DATA_BLOCK "DB1901_Config_Robots"   // DB1901
{ S7_Optimized_Access := 'FALSE' }
VERSION : 0.1
   VAR
      ReadWriteDeviceNo : Int := 1;
      CopyDeviceNO : Int := 0;
      Read : Bool := FALSE;
      Write : Bool := FALSE;
      Copy : Bool := FALSE;
      Config_Robots : Array[0..4] of Struct
         Type_Kuka : Bool;   // Kuka Robot
         Type_ABB : Bool;   // ABB Robot
         Type_Fanuc : Bool;   // Fanuc Robot
         Type_Motoman : Bool;   // Motoman (Yaskawa) Robot
         Type_5 : Bool;
         Type_6 : Bool;
         Type_7 : Bool;
         Type_8 : Bool;
         With_Shotware : Bool;   // Only ABB
         With_Tracking : Bool;
         With_Safetysoftware : Bool;   // EPS/Safemove or simmilar
         With_Synchronisation : Bool;   // EPS Sync switch, Breaktest, ...
         With_Testshot : Bool;   // With Test shot station
         With_Cleaning : Bool;   // With Cleaning (automaitc)
         With_Wet_Cleaning : Bool;   // With wet cleaning
         With_Wet_Cleaning_LFI : Bool;   // Water cleaning LFI
         With_Wet_Cleaning_Spray : Bool;   // Wet cleaning Spray
         With_IR_Station : Bool;   // With Infra red station
         With_Brush_Station : Bool;   // With Brush station (motor)
         With_Belt_Filter : Bool;   // With belt filter for LFI wet cleaning
         With_Air_Cleaner : Bool;   // With Air cleaning system for the mixinghead
         Spare_2_5 : Bool;
         Spare_2_6 : Bool;
         Spare_2_7 : Bool;
         MHNumber : Byte;
         InterfaceForTestShot : Byte;
         ForInterface : Array[1..16] of Bool;
      END_STRUCT;
   END_VAR
BEGIN
   Config_Robots[0].Type_Kuka := FALSE;
   Config_Robots[0].Type_ABB := FALSE;
   Config_Robots[0].Type_Fanuc := FALSE;
   Config_Robots[0].Type_Motoman := FALSE;
   Config_Robots[0].Type_5 := FALSE;
   Config_Robots[0].Type_6 := FALSE;
   Config_Robots[0].Type_7 := FALSE;
   Config_Robots[0].Type_8 := FALSE;
   Config_Robots[0].With_Shotware := FALSE;
   Config_Robots[0].With_Tracking := FALSE;
   Config_Robots[0].With_Safetysoftware := FALSE;
   Config_Robots[0].With_Synchronisation := TRUE;
   Config_Robots[0].With_Testshot := TRUE;
   Config_Robots[0].With_Cleaning := TRUE;
   Config_Robots[0].With_Wet_Cleaning := FALSE;
   Config_Robots[0].With_Wet_Cleaning_LFI := FALSE;
   Config_Robots[0].With_Wet_Cleaning_Spray := FALSE;
   Config_Robots[0].With_IR_Station := FALSE;
   Config_Robots[0].With_Brush_Station := FALSE;
   Config_Robots[0].With_Belt_Filter := FALSE;
   Config_Robots[0].With_Air_Cleaner := FALSE;
   Config_Robots[0].Spare_2_5 := FALSE;
   Config_Robots[0].Spare_2_6 := FALSE;
   Config_Robots[0].Spare_2_7 := FALSE;
   Config_Robots[1].Type_Kuka := FALSE;
   Config_Robots[1].Type_ABB := FALSE;
   Config_Robots[1].Type_Fanuc := FALSE;
   Config_Robots[1].Type_Motoman := FALSE;
   Config_Robots[1].Type_5 := FALSE;
   Config_Robots[1].Type_6 := FALSE;
   Config_Robots[1].Type_7 := FALSE;
   Config_Robots[1].Type_8 := FALSE;
   Config_Robots[1].With_Shotware := FALSE;
   Config_Robots[1].With_Tracking := FALSE;
   Config_Robots[1].With_Safetysoftware := FALSE;
   Config_Robots[1].With_Synchronisation := TRUE;
   Config_Robots[1].With_Testshot := TRUE;
   Config_Robots[1].With_Cleaning := TRUE;
   Config_Robots[1].With_Wet_Cleaning := FALSE;
   Config_Robots[1].With_Wet_Cleaning_LFI := FALSE;
   Config_Robots[1].With_Wet_Cleaning_Spray := FALSE;
   Config_Robots[1].With_IR_Station := FALSE;
   Config_Robots[1].With_Brush_Station := FALSE;
   Config_Robots[1].With_Belt_Filter := FALSE;
   Config_Robots[1].With_Air_Cleaner := FALSE;
   Config_Robots[1].Spare_2_5 := FALSE;
   Config_Robots[1].Spare_2_6 := FALSE;
   Config_Robots[1].Spare_2_7 := FALSE;
   Config_Robots[2].Type_Kuka := FALSE;
   Config_Robots[2].Type_ABB := FALSE;
   Config_Robots[2].Type_Fanuc := FALSE;
   Config_Robots[2].Type_Motoman := FALSE;
   Config_Robots[2].Type_5 := FALSE;
   Config_Robots[2].Type_6 := FALSE;
   Config_Robots[2].Type_7 := FALSE;
   Config_Robots[2].Type_8 := FALSE;
   Config_Robots[2].With_Shotware := FALSE;
   Config_Robots[2].With_Tracking := FALSE;
   Config_Robots[2].With_Safetysoftware := FALSE;
   Config_Robots[2].With_Synchronisation := FALSE;
   Config_Robots[2].With_Testshot := FALSE;
   Config_Robots[2].With_Cleaning := FALSE;
   Config_Robots[2].With_Wet_Cleaning := FALSE;
   Config_Robots[2].With_Wet_Cleaning_LFI := FALSE;
   Config_Robots[2].With_Wet_Cleaning_Spray := FALSE;
   Config_Robots[2].With_IR_Station := FALSE;
   Config_Robots[2].With_Brush_Station := FALSE;
   Config_Robots[2].With_Belt_Filter := FALSE;
   Config_Robots[2].With_Air_Cleaner := FALSE;
   Config_Robots[2].Spare_2_5 := FALSE;
   Config_Robots[2].Spare_2_6 := FALSE;
   Config_Robots[2].Spare_2_7 := FALSE;
   Config_Robots[3].Type_Kuka := FALSE;
   Config_Robots[3].Type_ABB := FALSE;
   Config_Robots[3].Type_Fanuc := FALSE;
   Config_Robots[3].Type_Motoman := FALSE;
   Config_Robots[3].Type_5 := FALSE;
   Config_Robots[3].Type_6 := FALSE;
   Config_Robots[3].Type_7 := FALSE;
   Config_Robots[3].Type_8 := FALSE;
   Config_Robots[3].With_Shotware := FALSE;
   Config_Robots[3].With_Tracking := FALSE;
   Config_Robots[3].With_Safetysoftware := FALSE;
   Config_Robots[3].With_Synchronisation := FALSE;
   Config_Robots[3].With_Testshot := FALSE;
   Config_Robots[3].With_Cleaning := FALSE;
   Config_Robots[3].With_Wet_Cleaning := FALSE;
   Config_Robots[3].With_Wet_Cleaning_LFI := FALSE;
   Config_Robots[3].With_Wet_Cleaning_Spray := FALSE;
   Config_Robots[3].With_IR_Station := FALSE;
   Config_Robots[3].With_Brush_Station := FALSE;
   Config_Robots[3].With_Belt_Filter := FALSE;
   Config_Robots[3].With_Air_Cleaner := FALSE;
   Config_Robots[3].Spare_2_5 := FALSE;
   Config_Robots[3].Spare_2_6 := FALSE;
   Config_Robots[3].Spare_2_7 := FALSE;
   Config_Robots[4].Type_Kuka := FALSE;
   Config_Robots[4].Type_ABB := FALSE;
   Config_Robots[4].Type_Fanuc := FALSE;
   Config_Robots[4].Type_Motoman := FALSE;
   Config_Robots[4].Type_5 := FALSE;
   Config_Robots[4].Type_6 := FALSE;
   Config_Robots[4].Type_7 := FALSE;
   Config_Robots[4].Type_8 := FALSE;
   Config_Robots[4].With_Shotware := FALSE;
   Config_Robots[4].With_Tracking := FALSE;
   Config_Robots[4].With_Safetysoftware := FALSE;
   Config_Robots[4].With_Synchronisation := FALSE;
   Config_Robots[4].With_Testshot := FALSE;
   Config_Robots[4].With_Cleaning := FALSE;
   Config_Robots[4].With_Wet_Cleaning := FALSE;
   Config_Robots[4].With_Wet_Cleaning_LFI := FALSE;
   Config_Robots[4].With_Wet_Cleaning_Spray := FALSE;
   Config_Robots[4].With_IR_Station := FALSE;
   Config_Robots[4].With_Brush_Station := FALSE;
   Config_Robots[4].With_Belt_Filter := FALSE;
   Config_Robots[4].With_Air_Cleaner := FALSE;
   Config_Robots[4].Spare_2_5 := FALSE;
   Config_Robots[4].Spare_2_6 := FALSE;
   Config_Robots[4].Spare_2_7 := FALSE;
   Config_Robots[1].ForInterface[1] := TRUE;
   Config_Robots[1].ForInterface[2] := TRUE;
   Config_Robots[1].ForInterface[3] := TRUE;
   Config_Robots[1].ForInterface[4] := TRUE;
   Config_Robots[1].ForInterface[5] := TRUE;
   Config_Robots[1].InterfaceForTestShot := 16#05;
   Config_Robots[0].MHNumber := 16#01;
   Config_Robots[0].InterfaceForTestShot := 16#05;
   Config_Robots[0].ForInterface[1] := TRUE;
   Config_Robots[0].ForInterface[2] := TRUE;
   Config_Robots[0].ForInterface[3] := TRUE;
   Config_Robots[0].ForInterface[4] := TRUE;
   Config_Robots[0].ForInterface[5] := TRUE;
   Config_Robots[0].ForInterface[6] := FALSE;
   Config_Robots[0].ForInterface[7] := FALSE;
   Config_Robots[0].ForInterface[8] := FALSE;
   Config_Robots[0].ForInterface[9] := FALSE;
   Config_Robots[0].ForInterface[10] := FALSE;
   Config_Robots[0].ForInterface[11] := FALSE;
   Config_Robots[0].ForInterface[12] := FALSE;
   Config_Robots[0].ForInterface[13] := FALSE;
   Config_Robots[0].ForInterface[14] := FALSE;
   Config_Robots[0].ForInterface[15] := FALSE;
   Config_Robots[0].ForInterface[16] := FALSE;
   Config_Robots[1].MHNumber := 16#01;
   Config_Robots[1].ForInterface[6] := FALSE;
   Config_Robots[1].ForInterface[7] := FALSE;
   Config_Robots[1].ForInterface[8] := FALSE;
   Config_Robots[1].ForInterface[9] := FALSE;
   Config_Robots[1].ForInterface[10] := FALSE;
   Config_Robots[1].ForInterface[11] := FALSE;
   Config_Robots[1].ForInterface[12] := FALSE;
   Config_Robots[1].ForInterface[13] := FALSE;
   Config_Robots[1].ForInterface[14] := FALSE;
   Config_Robots[1].ForInterface[15] := FALSE;
   Config_Robots[1].ForInterface[16] := FALSE;
   Config_Robots[2].MHNumber := 16#00;
   Config_Robots[2].InterfaceForTestShot := 16#00;
   Config_Robots[2].ForInterface[1] := FALSE;
   Config_Robots[2].ForInterface[2] := FALSE;
   Config_Robots[2].ForInterface[3] := FALSE;
   Config_Robots[2].ForInterface[4] := FALSE;
   Config_Robots[2].ForInterface[5] := FALSE;
   Config_Robots[2].ForInterface[6] := FALSE;
   Config_Robots[2].ForInterface[7] := FALSE;
   Config_Robots[2].ForInterface[8] := FALSE;
   Config_Robots[2].ForInterface[9] := FALSE;
   Config_Robots[2].ForInterface[10] := FALSE;
   Config_Robots[2].ForInterface[11] := FALSE;
   Config_Robots[2].ForInterface[12] := FALSE;
   Config_Robots[2].ForInterface[13] := FALSE;
   Config_Robots[2].ForInterface[14] := FALSE;
   Config_Robots[2].ForInterface[15] := FALSE;
   Config_Robots[2].ForInterface[16] := FALSE;
   Config_Robots[3].MHNumber := 16#00;
   Config_Robots[3].InterfaceForTestShot := 16#00;
   Config_Robots[3].ForInterface[1] := FALSE;
   Config_Robots[3].ForInterface[2] := FALSE;
   Config_Robots[3].ForInterface[3] := FALSE;
   Config_Robots[3].ForInterface[4] := FALSE;
   Config_Robots[3].ForInterface[5] := FALSE;
   Config_Robots[3].ForInterface[6] := FALSE;
   Config_Robots[3].ForInterface[7] := FALSE;
   Config_Robots[3].ForInterface[8] := FALSE;
   Config_Robots[3].ForInterface[9] := FALSE;
   Config_Robots[3].ForInterface[10] := FALSE;
   Config_Robots[3].ForInterface[11] := FALSE;
   Config_Robots[3].ForInterface[12] := FALSE;
   Config_Robots[3].ForInterface[13] := FALSE;
   Config_Robots[3].ForInterface[14] := FALSE;
   Config_Robots[3].ForInterface[15] := FALSE;
   Config_Robots[3].ForInterface[16] := FALSE;
   Config_Robots[4].MHNumber := 16#00;
   Config_Robots[4].InterfaceForTestShot := 16#00;
   Config_Robots[4].ForInterface[1] := FALSE;
   Config_Robots[4].ForInterface[2] := FALSE;
   Config_Robots[4].ForInterface[3] := FALSE;
   Config_Robots[4].ForInterface[4] := FALSE;
   Config_Robots[4].ForInterface[5] := FALSE;
   Config_Robots[4].ForInterface[6] := FALSE;
   // 10 more start values not shown
END_DATA_BLOCK

DATA_BLOCK "GetToolShotValues_DB"   // DB1930
{ S7_Optimized_Access := 'FALSE' }
VERSION : 0.1
"GetToolShotValues"
BEGIN
   IN_MachineNo := 1;
   IN_EnableTool := TRUE;
END_DATA_BLOCK

DATA_BLOCK "FB1931_ToolAllocationList_DB"   // DB1931
{ S7_Optimized_Access := 'TRUE' }
VERSION : 0.1
"FB1931_ToolAllocationList"
BEGIN
END_DATA_BLOCK

DATA_BLOCK "DB2000_FRA<->KM"   // DB2000
{ S7_Optimized_Access := 'FALSE' }
VERSION : 0.1
   VAR
      AP_Shottime : Int := 0;   // Schusszeit in ms
      AP_MVH : Int := 0;   // Mischungsverhältnis in 0,1%
      AP_Weight : Int := 0;   // Gesamtgewicht pro Sekunde in 0,1 Gramm
      FRA1_Stat : "UDT2000_KM_FRA";
      FRA1_PrgNr : Byte := B#16#0;
      Bit_FT1_sel : Bool := FALSE;
      Bit_FRA1_Sel : Bool := FALSE;
      TS1_Offset : Byte := B#16#0;
      Input : "UDT2001_Input_Faurecia";
      Output : "UDT2002_Output_Faurecia";
   END_VAR
BEGIN
END_DATA_BLOCK

DATA_BLOCK "PN_Devices"   // DB2023
{ S7_Optimized_Access := 'TRUE' }
VERSION : 0.1
   VAR
      LADDR : Hw_IoSystem := 257;
      MODE : UInt := 4;
      RETVAL : Int;
      Device_available : Array[0..1023] of Bool;
   END_VAR
BEGIN
   // Device_available[2] : pn-mixhead
   // Device_available[1] : pn-flow1
   // Device_available[0] : Bei mindestens einem der IO-Devices liegt eine Störung vor.
END_DATA_BLOCK

DATA_BLOCK "PB_Devices"   // DB2024
{ S7_Optimized_Access := 'TRUE' }
VERSION : 0.1
   VAR
      LADDR : Hw_IoSystem := 296;
      MODE : UInt := 4;
      RETVAL : Int;
      Device_available : Array[0..127] of Bool;
   END_VAR
BEGIN
END_DATA_BLOCK

// folder: System blocks/Program resources

DATA_BLOCK "DB55_Temp_HD_WT_MK1_K1"   // DB55
{ S7_Optimized_Access := 'TRUE' }
AUTHOR : Simatic
FAMILY : IEC
NAME : IEC_TMR
VERSION : 1.0
"IEC_TIMER"
BEGIN
END_DATA_BLOCK

DATA_BLOCK "DB56_Temp_HD_WT_MK1_K2"   // DB56
{ S7_Optimized_Access := 'TRUE' }
AUTHOR : Simatic
FAMILY : IEC
NAME : IEC_TMR
VERSION : 1.0
"IEC_TIMER"
BEGIN
END_DATA_BLOCK

DATA_BLOCK "DB60_Temp_ND_WT_MK1_K1"   // DB60
{ S7_Optimized_Access := 'TRUE' }
AUTHOR : Simatic
FAMILY : IEC
NAME : IEC_TMR
VERSION : 1.0
"IEC_TIMER"
BEGIN
END_DATA_BLOCK

DATA_BLOCK "DB61_Temp_ND_WT_MK1_K2"   // DB61
{ S7_Optimized_Access := 'TRUE' }
AUTHOR : Simatic
FAMILY : IEC
NAME : IEC_TMR
VERSION : 1.0
"IEC_TIMER"
BEGIN
END_DATA_BLOCK

// folder: (top level)

FUNCTION_BLOCK "FB_MouldEditor_HMI"   // FB4, SCL
{ S7_Optimized_Access := 'FALSE' }
VERSION : 0.1
   VAR_INPUT
      INiAmountMeteringUnits : Int;   // Amount of metering units
   END_VAR
   VAR_IN_OUT
      IOuMouldEditor_HMI : "typeMouldEditor_HMI";   // Data of mould editor - actual
   END_VAR
   VAR
      SuMouldEditor_HMI : "typeMouldEditor_HMI";   // Data of mould editor - last PLC cycle
   END_VAR
   VAR_TEMP
      TiPartShotAmount : Int;   // Amount of part shoots at this tool
      TiComponentAmount : Int;   // Amount of components at this part shot (depending on MH no)
      TiLoop_PS : Int;   // Value for loop - partial shot number
      TiLoop : Int;   // Value for loop - general
      TiLoop_Flow : Int;   // Value for loop - flow
      TiLoop_Ratio : Int;   // Value for loop - ratio
      OUTrSumFlow : Real;
      RefComp : Int;
      TrFlowRefComp : Real;
      MouldNo : Int;
      OUTrSumRatio : Real;
      OUTrDifRatio : Real;
      OUTrDifTotalFlow : Real;
      TrMaxTotalFlow : Real;
      Nullbyte : Byte;
      Retval : Int;
      Ti_alloc_list : Int;
   END_VAR
BEGIN

   IF "TP-Bereichszeiger".Picturenumber.Bildnummer = 892 THEN   //  Screen no. of editor mould foaming data
       //_________________________________________________________________________________    
       // Decleration of part shots and shot amount
       "InterfaceVisu".AmountTools := "AmountTools";
       "InterfaceVisu".AmountAlloactionAutomatic := "AmountAllocationAutomatic"; //<-- Array value of allocation places (default 200)
       "InterfaceVisu".AmountPartShots := "AmountPartShots"; //<-- Array value of part shots (default 8)
       //_________________________________________________________________________________    
       //  Limit values
       #IOuMouldEditor_HMI.sSelected.iTool := LIMIT(MN := 1, IN := #IOuMouldEditor_HMI.sSelected.iTool, MX := "InterfaceVisu".AmountTools);
       #IOuMouldEditor_HMI.sSelected.sPS.iPS := LIMIT(MN := 0, IN := #IOuMouldEditor_HMI.sSelected.sPS.iPS, MX := "AmountPartShots");
       //_________________________________________________________________________________    
       // Part shot increase
       IF #IOuMouldEditor_HMI.sStatusBits.xPartShotAmount_increase THEN
           #IOuMouldEditor_HMI.sStatusBits.xPartShotAmount_increase := False;
           IF #IOuMouldEditor_HMI.uTools.PartShot_Amount < "AmountPartShots" THEN
               #IOuMouldEditor_HMI.uTools.PartShot_Amount := #IOuMouldEditor_HMI.uTools.PartShot_Amount + 1;
           END_IF;
       END_IF;
       // Part shot decrease
       IF #IOuMouldEditor_HMI.sStatusBits.xPartShotAmount_decrease THEN
           #IOuMouldEditor_HMI.sStatusBits.xPartShotAmount_decrease := False;
           IF #IOuMouldEditor_HMI.uTools.PartShot_Amount > 0 THEN
               #IOuMouldEditor_HMI.uTools.PartShot_Amount := #IOuMouldEditor_HMI.uTools.PartShot_Amount - 1;
           END_IF;
       END_IF;
       //_________________________________________________________________________________    
       // Last part shot / last tool selected
       "InterfaceVisu".LastPartShot := #IOuMouldEditor_HMI.uTools.PartShot_Amount >= "AmountPartShots";
       "InterfaceVisu".LastTool := #IOuMouldEditor_HMI.sSelected.iTool >= "InterfaceVisu".AmountTools;
       //_________________________________________________________________________________    
       // Shot time from s5time to real
       "InterfaceVisu".MaxShottime := DINT_TO_REAL(TIME_TO_DINT(S5TIME_TO_TIME("DB700_Machine".Machine[1].Max_ShotTime)))/1000;
       "InterfaceVisu".MinShottime := DINT_TO_REAL(TIME_TO_DINT(S5TIME_TO_TIME("DB700_Machine".Machine[1].Min_ShotTime)))/1000;
       //_________________________________________________________________________________    
       // Diverse Abarbeitungen für die Anzeige des Schäumprograms    
       REGION 1. Herusfinden der Komponenten- Anzahl an dem ausgewählten Mischkopf
           #TiComponentAmount := "DB704_MH_Value".Mixinghead[#IOuMouldEditor_HMI.arShotSet[#IOuMouldEditor_HMI.sSelected.sPS.iPS].MHNo].AmountComponent;
       END_REGION
       #RefComp := LIMIT(MN := 1, IN := #IOuMouldEditor_HMI.sSelected.sPS.RefComponent, MX := #TiComponentAmount);
       REGION 2. Anzeigen der Komponenten- Namen je zugeordneten Mischkopf im Schäumprogramm
           // Max Flow for limits
           // Component used at this mixinghead
           // 2 Point at this mixinghead
           IF #IOuMouldEditor_HMI.sSelected.sPS.iPS <> 0 THEN
               FOR #TiLoop_Flow := 1 TO #TiComponentAmount DO
                   "InterfaceVisu".NameComp[#TiLoop_Flow] := "DB614_MH_State".MH_Connection[#IOuMouldEditor_HMI.arShotSet[#IOuMouldEditor_HMI.sSelected.sPS.iPS].MHNo].Name[#TiLoop_Flow];
                   // Max flow for all components = 0 if Refcomponent and selected refcomp is 0
                   IF #IOuMouldEditor_HMI.sSelected.sPS.arFlow[#RefComp] = 0 THEN
                       // all limits to 0 excluding the ref component
                       "InterfaceVisu".MaxFlow[#TiLoop_Flow] := 0;
                       "InterfaceVisu".MaxFlow[#RefComp] := "DB614_MH_State".MH_Connection[#IOuMouldEditor_HMI.arShotSet[#IOuMouldEditor_HMI.sSelected.sPS.iPS].MHNo].MaxFlow[#RefComp];
                   ELSE
                       "InterfaceVisu".MaxFlow[#TiLoop_Flow] := "DB614_MH_State".MH_Connection[#IOuMouldEditor_HMI.arShotSet[#IOuMouldEditor_HMI.sSelected.sPS.iPS].MHNo].MaxFlow[#TiLoop_Flow];
                   END_IF;
                   // Min flow = 0 if MR = 0 at this component
                   IF #IOuMouldEditor_HMI.sSelected.sPS.arRatio[#TiLoop_Flow] = 0 THEN
                       "InterfaceVisu".MinFlow[#TiLoop_Flow] := 0;
                   ELSE
                       "InterfaceVisu".MinFlow[#TiLoop_Flow] := "DB614_MH_State".MH_Connection[#IOuMouldEditor_HMI.arShotSet[#IOuMouldEditor_HMI.sSelected.sPS.iPS].MHNo].MinFlow[#TiLoop_Flow];
                   END_IF;

                   "InterfaceVisu".CompAtMixinghead[#TiLoop_Flow] := True;
                   //"InterfaceVisu"."2PoinMovementComp"[#TiLoop_Flow] := "DB753_MeteringPump".Pump["DB704_MH_Value".Mixinghead["DB925_ShotData".Tool[#IOuMouldEditor_HMI.sSelected.iTool].Shot[#IOuMouldEditor_HMI.sSelected.sPS.iPS].MHNo].MH_Connection[#TiLoop_Flow].Pump_No].With_2Point;
               END_FOR;
               // Set not used components to "0"
               IF #TiComponentAmount < 6 THEN
                   FOR #TiLoop_Flow := #TiComponentAmount + 1 TO 6 DO
                       "InterfaceVisu".CompAtMixinghead[#TiLoop_Flow] := FALSE;
                       "InterfaceVisu"."2PoinMovementComp"[#TiLoop_Flow] := False;
                       "InterfaceVisu".MinFlow[#TiLoop_Flow] := 0;
                       "InterfaceVisu".MaxFlow[#TiLoop_Flow] := 0;
                       "InterfaceVisu".NameComp[#TiLoop_Flow] := '   ';
                   END_FOR;
               END_IF;
           END_IF;
       END_REGION
       REGION 3. Calculate max total flow
           // Check for each part shot the MH number and the amount of components
           FOR #TiLoop_PS := 1 TO "AmountPartShots" DO
               #TrMaxTotalFlow := 0;
               FOR #TiLoop := 1 TO BYTE_TO_INT("DB704_MH_Value".Mixinghead[#IOuMouldEditor_HMI.arShotSet[#TiLoop_PS].MHNo].AmountComponent) DO
                   // Max total flow
                   #TrMaxTotalFlow := #TrMaxTotalFlow +
                   "DB614_MH_State".MH_Connection[#IOuMouldEditor_HMI.arShotSet[#TiLoop_PS].MHNo].MaxFlow[#TiLoop];
               END_FOR;
               "InterfaceVisu".MaxTotalFlow[#TiLoop_PS] := #TrMaxTotalFlow;
           END_FOR;
           //#IOuMouldEditor_HMI.sCalculatedValues.arTotalFlow[#IOuMouldEditor_HMI.sSelected.sPS.iPS] := LIMIT(MN := 0, IN := #IOuMouldEditor_HMI.sCalculatedValues.arTotalFlow[#IOuMouldEditor_HMI.sSelected.sPS.iPS], MX := "InterfaceVisu".MaxTotalFlow[#IOuMouldEditor_HMI.sSelected.sPS.iPS]);
       END_REGION
       REGION 4. Übernehmen der Hochdruck- Kreislaufwerte an dem Mischkopf der in dem Teilschuß eingetragen wurde
           IF "InterfaceVisu".SetHDValue = True THEN
               // Mixinghead No. set by Shot Data (classic)    
               IF "DB790_PlantParameter".Bit.MHNofromInterface = False THEN
                   FOR #TiLoop_Flow := 1 TO #TiComponentAmount DO
                       // If a component is "0" don't write it to the HP values
                       IF "DB925_ShotData_1".Tool[#IOuMouldEditor_HMI.sSelected.iTool].Shot[#IOuMouldEditor_HMI.sSelected.sPS.iPS].Flow[#TiLoop_Flow] <> 0 THEN
                           "DB704_MH_Value".Mixinghead["DB925_ShotData_1".Tool[#IOuMouldEditor_HMI.sSelected.iTool].Shot[#IOuMouldEditor_HMI.sSelected.sPS.iPS].MHNo].MH_Connection[#TiLoop_Flow].Flow_HP_Circ :=
                           "DB925_ShotData_1".Tool[#IOuMouldEditor_HMI.sSelected.iTool].Shot[#IOuMouldEditor_HMI.sSelected.sPS.iPS].Flow[#TiLoop_Flow];
                       END_IF;
                   END_FOR;

                   // Mixinghead No. set by Interface
               ELSIF "DB790_PlantParameter".Bit.MHNofromInterface = true THEN
                   // If Mixinghead number is set bei Interface, check if selected program is allocated, tool is installed, and then write HP values to right mixinghead
                   FOR #TiLoop := 1 TO "DB790_PlantParameter".AmountToolStation DO  // Check all Tool codes at all interfaces
                       #MouldNo := "DB005_RS<->Extern".MC_Interface[#TiLoop].Data_from_MC.Toolcode;
                       IF "DB940_Tool_alloc_automatic".Alloc_stationTool[#MouldNo] = "DB925_ShotData_1".Tool_No THEN    // compare if selected tool match with one of the interfaces
                           FOR #TiLoop_Flow := 1 TO #TiComponentAmount DO
                               // If a component is "0" don't write it to the HP values
                               IF "DB925_ShotData_1".Tool[#IOuMouldEditor_HMI.sSelected.iTool].Shot[#IOuMouldEditor_HMI.sSelected.sPS.iPS].Flow[#TiLoop_Flow] <> 0 THEN
                                   "DB704_MH_Value".Mixinghead[#TiLoop].MH_Connection[#TiLoop_Flow].Flow_HP_Circ := "DB925_ShotData_1".Tool[#IOuMouldEditor_HMI.sSelected.iTool].Shot[#IOuMouldEditor_HMI.sSelected.sPS.iPS].Flow[#TiLoop_Flow];
                               END_IF;
                           END_FOR;
                       ELSE // If tool is not allocated ask where to copy the HP values

                           IF "InterfaceVisu".PopUp_MH_No = true THEN
                               FOR #TiLoop_Flow := 1 TO #TiComponentAmount DO
                                   // If a component is "0" don't write it to the HP values
                                   IF "DB925_ShotData_1".Tool[#IOuMouldEditor_HMI.sSelected.iTool].Shot[#IOuMouldEditor_HMI.sSelected.sPS.iPS].Flow[#TiLoop_Flow] <> 0 THEN
                                       "DB704_MH_Value".Mixinghead["InterfaceVisu".MH_No_for_HPValues].MH_Connection[#TiLoop_Flow].Flow_HP_Circ := "DB925_ShotData_1".Tool[#IOuMouldEditor_HMI.sSelected.iTool].Shot[#IOuMouldEditor_HMI.sSelected.sPS.iPS].Flow[#TiLoop_Flow];
                                   END_IF;
                                   "InterfaceVisu".PopUp_MH_No := false;   // Pop up: Write HP values to selected mixinghead
                               END_FOR;
                           ELSIF "InterfaceVisu".HPValuesSet = false AND #TiLoop >= "DB790_PlantParameter".AmountToolStation THEN
                               "InterfaceVisu".PopUp_MH_No := True;   // Pop up: Write HP values to selected mixinghead
                           END_IF;
                       END_IF;
                   END_FOR;
               END_IF;

               "InterfaceVisu".SetHDValue := 0;
           END_IF;
       END_REGION
       REGION 5. Check HP values
       FOR #TiLoop_Flow := 1 TO #TiComponentAmount DO
           IF REAL_TO_DINT("DB704_MH_Value".Mixinghead[#IOuMouldEditor_HMI.arShotSet[#IOuMouldEditor_HMI.sSelected.sPS.iPS].MHNo].MH_Connection[#TiLoop_Flow].Flow_HP_Circ) =
               REAL_TO_DINT(#IOuMouldEditor_HMI.arShotSet[#IOuMouldEditor_HMI.sSelected.sPS.iPS].Flow[#TiLoop_Flow]) OR
               REAL_TO_DINT(#IOuMouldEditor_HMI.arShotSet[#IOuMouldEditor_HMI.sSelected.sPS.iPS].Flow[#TiLoop_Flow]) = 0 THEN
               "InterfaceVisu".HPValuesSet := TRUE;
           ELSE
               "InterfaceVisu".HPValuesSet := FALSE;
               EXIT;
           END_IF;
       END_FOR;
       END_REGION
       //_________________________________________________________________________________    
       REGION Limit MR/Pressure
           FOR #TiLoop_Ratio := 1 TO 6 DO
               #IOuMouldEditor_HMI.sSelected.sPS.arRatio[#TiLoop_Ratio] := LIMIT(MN := 0, IN := #IOuMouldEditor_HMI.sSelected.sPS.arRatio[#TiLoop_Ratio], MX := 999999999);
               #IOuMouldEditor_HMI.sSelected.sPS.arPressure[#TiLoop_Ratio] := LIMIT(MN := 0, IN := #IOuMouldEditor_HMI.sSelected.sPS.arPressure[#TiLoop_Ratio], MX := 2500);
           END_FOR;
       END_REGION
       #TiPartShotAmount := #IOuMouldEditor_HMI.uTools.PartShot_Amount;
       #TiPartShotAmount := LIMIT(MN := 0, IN := #TiPartShotAmount, MX := "AmountPartShots");
       //_________________________________________________________________________________    
       REGION Tool number changed -> copy all data
           IF #IOuMouldEditor_HMI.sSelected.iTool <> #SuMouldEditor_HMI.sSelected.iTool OR #IOuMouldEditor_HMI.sStatusBits.xDiscardChanges THEN

               #IOuMouldEditor_HMI.sStatusBits.xValueChanged := FALSE;
               #IOuMouldEditor_HMI.sStatusBits.xSafeChanges := FALSE;
               #IOuMouldEditor_HMI.sStatusBits.xDiscardChanges := FALSE;

               FOR #TiLoop_PS := 1 TO "AmountPartShots" DO
                   // When the selected Tool less or equal 100 is, take the values from DB925
                   IF #IOuMouldEditor_HMI.sSelected.iTool <= "AmountToolsDB" THEN
                       #IOuMouldEditor_HMI.arShotSet[#TiLoop_PS] := "DB925_ShotData_1".Tool[#IOuMouldEditor_HMI.sSelected.iTool].Shot[#TiLoop_PS];
                   END_IF;
                   // When the selected Tool bigger than 100 and less or equal 200 is, take the values from DB926
                   IF #IOuMouldEditor_HMI.sSelected.iTool > "AmountToolsDB" AND #IOuMouldEditor_HMI.sSelected.iTool <= (2*"AmountToolsDB") THEN
                       #IOuMouldEditor_HMI.arShotSet[#TiLoop_PS] := "DB926_ShotData_2".Tool[#IOuMouldEditor_HMI.sSelected.iTool-"AmountToolsDB"].Shot[#TiLoop_PS];
                   END_IF;
               END_FOR;

               // For some reason it is not possible to copy the flow consumption in the loop befor
               FOR #TiLoop_PS := 1 TO "AmountPartShots" DO
                   // SumFlow
                   #OUTrSumFlow := 0;

                   FOR #TiLoop_Flow := 1 TO 6 DO
                       #OUTrSumFlow := #OUTrSumFlow + #IOuMouldEditor_HMI.arShotSet[#TiLoop_PS].Flow[#TiLoop_Flow];
                   END_FOR;
                   #IOuMouldEditor_HMI.sCalculatedValues.arTotalFlow[#TiLoop_PS] := #OUTrSumFlow;
               END_FOR;

               #IOuMouldEditor_HMI.uTools := "DB930_Tools".Tool[#IOuMouldEditor_HMI.sSelected.iTool];

               //  Selected - partial shot
               #IOuMouldEditor_HMI.sSelected.sPS.iPS := 1;

               FOR #TiLoop := 1 TO #TiComponentAmount DO
                   #IOuMouldEditor_HMI.sSelected.sPS.arFlow[#TiLoop] := #IOuMouldEditor_HMI.arShotSet[1].Flow[#TiLoop];
                   #IOuMouldEditor_HMI.sSelected.sPS.arPressure[#TiLoop] := #IOuMouldEditor_HMI.arShotSet[1].Pressure[#TiLoop];
               END_FOR;

               // ----
               //  Save data for the last cycle to recognize changes of the values
               #SuMouldEditor_HMI := #IOuMouldEditor_HMI;
               // ----

           END_IF;
       END_REGION
       //_________________________________________________________________________________    
       REGION Tool name changed
           IF #IOuMouldEditor_HMI.uTools.tool_name <> #SuMouldEditor_HMI.uTools.tool_name THEN
           // ----
           //  Save data for the last cycle to recognize changes of the values
           #IOuMouldEditor_HMI.sStatusBits.xValueChanged := TRUE;
           #SuMouldEditor_HMI := #IOuMouldEditor_HMI;
           // ----
           END_IF;
       END_REGION
       //_________________________________________________________________________________    
       REGION Partialshot number increase -> fill partialshot with meaningful values
           IF #IOuMouldEditor_HMI.uTools.PartShot_Amount > #SuMouldEditor_HMI.uTools.PartShot_Amount THEN

               #IOuMouldEditor_HMI.sSelected.sPS.iPS := #IOuMouldEditor_HMI.uTools.PartShot_Amount;

               // First part shot use default values
               IF #IOuMouldEditor_HMI.uTools.PartShot_Amount = 1 THEN

                   #IOuMouldEditor_HMI.uTools.EnableTool := 1;
                   #IOuMouldEditor_HMI.arShotSet[#IOuMouldEditor_HMI.sSelected.sPS.iPS].MHNo := 1;
                   #IOuMouldEditor_HMI.arShotSet[#IOuMouldEditor_HMI.sSelected.sPS.iPS].FoamingTime := 1.00;
                   #IOuMouldEditor_HMI.arShotSet[#IOuMouldEditor_HMI.sSelected.sPS.iPS].PartWeight := 100.00;

                   FOR #TiLoop := 1 TO 6 DO
                       #IOuMouldEditor_HMI.arShotSet[#IOuMouldEditor_HMI.sSelected.sPS.iPS].Pressure[#TiLoop] := 0;
                   END_FOR;

                   #IOuMouldEditor_HMI.arShotSet[#IOuMouldEditor_HMI.sSelected.sPS.iPS].Flow[1] := 100.00;
                   FOR #TiLoop := 2 TO 6 DO
                       #IOuMouldEditor_HMI.arShotSet[#IOuMouldEditor_HMI.sSelected.sPS.iPS].Flow[#TiLoop] := 0;
                   END_FOR;
                   #IOuMouldEditor_HMI.arShotSet[#IOuMouldEditor_HMI.sSelected.sPS.iPS].RefComponent := 1;

               ELSE // Second and following part shots values from part shot befor
                   #IOuMouldEditor_HMI.arShotSet[#IOuMouldEditor_HMI.sSelected.sPS.iPS].MHNo := #IOuMouldEditor_HMI.arShotSet[#IOuMouldEditor_HMI.sSelected.sPS.iPS - 1].MHNo;
                   #IOuMouldEditor_HMI.arShotSet[#IOuMouldEditor_HMI.sSelected.sPS.iPS].FoamingTime := #IOuMouldEditor_HMI.arShotSet[#IOuMouldEditor_HMI.sSelected.sPS.iPS - 1].FoamingTime;
                   #IOuMouldEditor_HMI.arShotSet[#IOuMouldEditor_HMI.sSelected.sPS.iPS].PartWeight := #IOuMouldEditor_HMI.arShotSet[#IOuMouldEditor_HMI.sSelected.sPS.iPS - 1].PartWeight;
                   #IOuMouldEditor_HMI.arShotSet[#IOuMouldEditor_HMI.sSelected.sPS.iPS].PartShotDisable := #IOuMouldEditor_HMI.arShotSet[#IOuMouldEditor_HMI.sSelected.sPS.iPS - 1].PartShotDisable;
                   #IOuMouldEditor_HMI.arShotSet[#IOuMouldEditor_HMI.sSelected.sPS.iPS].CPMoveAfterShot := #IOuMouldEditor_HMI.arShotSet[#IOuMouldEditor_HMI.sSelected.sPS.iPS - 1].CPMoveAfterShot;
                   #IOuMouldEditor_HMI.arShotSet[#IOuMouldEditor_HMI.sSelected.sPS.iPS].PartCounter := #IOuMouldEditor_HMI.arShotSet[#IOuMouldEditor_HMI.sSelected.sPS.iPS - 1].PartCounter;
                   #IOuMouldEditor_HMI.arShotSet[#IOuMouldEditor_HMI.sSelected.sPS.iPS].PurgeMHAfterShot := #IOuMouldEditor_HMI.arShotSet[#IOuMouldEditor_HMI.sSelected.sPS.iPS - 1].PurgeMHAfterShot;

                   FOR #TiLoop := 1 TO 6 DO
                       #IOuMouldEditor_HMI.arShotSet[#IOuMouldEditor_HMI.sSelected.sPS.iPS].Pressure[#TiLoop] := #IOuMouldEditor_HMI.arShotSet[#IOuMouldEditor_HMI.sSelected.sPS.iPS - 1].Pressure[#TiLoop];
                       #IOuMouldEditor_HMI.arShotSet[#IOuMouldEditor_HMI.sSelected.sPS.iPS].Flow[#TiLoop] := #IOuMouldEditor_HMI.arShotSet[#IOuMouldEditor_HMI.sSelected.sPS.iPS - 1].Flow[#TiLoop];
                   END_FOR;
                   #IOuMouldEditor_HMI.arShotSet[#IOuMouldEditor_HMI.sSelected.sPS.iPS].RefComponent := #IOuMouldEditor_HMI.arShotSet[#IOuMouldEditor_HMI.sSelected.sPS.iPS - 1].RefComponent;

               END_IF;

               // SumFlow
               #OUTrSumFlow := 0;

               FOR #TiLoop_Flow := 1 TO 6 DO
                   #OUTrSumFlow := #OUTrSumFlow + #IOuMouldEditor_HMI.arShotSet[#IOuMouldEditor_HMI.sSelected.sPS.iPS].Flow[#TiLoop_Flow];
               END_FOR;
               #IOuMouldEditor_HMI.sCalculatedValues.arTotalFlow[#IOuMouldEditor_HMI.sSelected.sPS.iPS] := #OUTrSumFlow;

               //  Selected partial shot
               FOR #TiLoop := 1 TO 6 DO
                   #IOuMouldEditor_HMI.sSelected.sPS.arFlow[#TiLoop] := #IOuMouldEditor_HMI.arShotSet[#IOuMouldEditor_HMI.sSelected.sPS.iPS].Flow[#TiLoop];
                   #IOuMouldEditor_HMI.sSelected.sPS.arPressure[#TiLoop] := #IOuMouldEditor_HMI.arShotSet[#IOuMouldEditor_HMI.sSelected.sPS.iPS].Pressure[#TiLoop];
               END_FOR;
               #IOuMouldEditor_HMI.sSelected.sPS.arRatio[1] := 100.00;
               FOR #TiLoop := 2 TO 6 DO
                   #IOuMouldEditor_HMI.sSelected.sPS.arRatio[#TiLoop] := 0;
               END_FOR;
               // ----
               // Set max total flow once to avoid tolerance alarm
               "InterfaceVisu".MaxTotalFlow[#IOuMouldEditor_HMI.sSelected.sPS.iPS] := #IOuMouldEditor_HMI.sCalculatedValues.arTotalFlow[#IOuMouldEditor_HMI.sSelected.sPS.iPS];
               //  Value changed + Save data for the last cycle to recognize changes of the values
               #IOuMouldEditor_HMI.sStatusBits.xValueChanged := TRUE;
               #SuMouldEditor_HMI := #IOuMouldEditor_HMI;
               // ----
           END_IF;
       END_REGION
       //_________________________________________________________________________________    
       REGION Partialshot number decrease -> fill partialshot with 0
           IF #IOuMouldEditor_HMI.uTools.PartShot_Amount < #SuMouldEditor_HMI.uTools.PartShot_Amount THEN

               #IOuMouldEditor_HMI.sSelected.sPS.iPS := #IOuMouldEditor_HMI.uTools.PartShot_Amount;

               // Reset all part shot values after the last used part shot
               FOR #TiLoop_PS := BYTE_TO_INT(#IOuMouldEditor_HMI.uTools.PartShot_Amount) + 1 TO "AmountPartShots" DO
                   #IOuMouldEditor_HMI.arShotSet[#TiLoop_PS].MHNo := 0;
                   #IOuMouldEditor_HMI.arShotSet[#TiLoop_PS].FoamingTime := 0;
                   #IOuMouldEditor_HMI.arShotSet[#TiLoop_PS].PartWeight := 0;
                   #IOuMouldEditor_HMI.arShotSet[#TiLoop_PS].PartShotDisable := 0;
                   #IOuMouldEditor_HMI.arShotSet[#TiLoop_PS].CPMoveAfterShot := 0;
                   #IOuMouldEditor_HMI.arShotSet[#TiLoop_PS].PartCounter := 0;
                   #IOuMouldEditor_HMI.arShotSet[#TiLoop_PS].PurgeMHAfterShot := 0;

                   FOR #TiLoop := 1 TO 6 DO
                       #IOuMouldEditor_HMI.arShotSet[#TiLoop_PS].Pressure[#TiLoop] := 0;
                   END_FOR;

                   FOR #TiLoop := 1 TO 6 DO
                       #IOuMouldEditor_HMI.arShotSet[#TiLoop_PS].Flow[#TiLoop] := 0;
                   END_FOR;
                   #IOuMouldEditor_HMI.arShotSet[#TiLoop_PS].RefComponent := 1;
               END_FOR;

               //  Value changed + Save data for the last cycle to recognize changes of the values
               #IOuMouldEditor_HMI.sStatusBits.xValueChanged := TRUE;
               #SuMouldEditor_HMI := #IOuMouldEditor_HMI;
               // ----

           END_IF;
       END_REGION
       //_________________________________________________________________________________    
       REGION Partialshot number - changed
           IF #IOuMouldEditor_HMI.sSelected.sPS.iPS <> #SuMouldEditor_HMI.sSelected.sPS.iPS THEN
               FOR #TiLoop := 1 TO #TiComponentAmount DO
                   #IOuMouldEditor_HMI.sSelected.sPS.arFlow[#TiLoop] := #IOuMouldEditor_HMI.arShotSet[#IOuMouldEditor_HMI.sSelected.sPS.iPS].Flow[#TiLoop];
                   #IOuMouldEditor_HMI.sSelected.sPS.arPressure[#TiLoop] := #IOuMouldEditor_HMI.arShotSet[#IOuMouldEditor_HMI.sSelected.sPS.iPS].Pressure[#TiLoop];
               END_FOR;

               #IOuMouldEditor_HMI.sSelected.sPS.RefComponent := #IOuMouldEditor_HMI.arShotSet[#IOuMouldEditor_HMI.sSelected.sPS.iPS].RefComponent;
               // Values 2-point adjust
               // #IOuMouldEditor_HMI.sSelected.sPS."2PoinMovement_Comp01" := #IOuMouldEditor_HMI.arShotSet[#IOuMouldEditor_HMI.sSelected.sPS.iPS]."2PoinMovement_Comp01";
               // #IOuMouldEditor_HMI.sSelected.sPS."2PoinMovement_Comp02" := #IOuMouldEditor_HMI.arShotSet[#IOuMouldEditor_HMI.sSelected.sPS.iPS]."2PoinMovement_Comp02";
               // #IOuMouldEditor_HMI.sSelected.sPS."2PoinMovement_Comp03" := #IOuMouldEditor_HMI.arShotSet[#IOuMouldEditor_HMI.sSelected.sPS.iPS]."2PoinMovement_Comp03";
               // #IOuMouldEditor_HMI.sSelected.sPS."2PoinMovement_Comp04" := #IOuMouldEditor_HMI.arShotSet[#IOuMouldEditor_HMI.sSelected.sPS.iPS]."2PoinMovement_Comp04";
               // #IOuMouldEditor_HMI.sSelected.sPS."2PoinMovement_Comp05" := #IOuMouldEditor_HMI.arShotSet[#IOuMouldEditor_HMI.sSelected.sPS.iPS]."2PoinMovement_Comp05";
               // #IOuMouldEditor_HMI.sSelected.sPS."2PoinMovement_Comp06" := #IOuMouldEditor_HMI.arShotSet[#IOuMouldEditor_HMI.sSelected.sPS.iPS]."2PoinMovement_Comp06";

               //------------------------------------------------------------------------------------------------------------------------------------------------
               // Reference component = 100%
               #RefComp := LIMIT(MN := 1, IN := #IOuMouldEditor_HMI.sSelected.sPS.RefComponent, MX := #TiComponentAmount);
               #IOuMouldEditor_HMI.sSelected.sPS.RefComponent := #RefComp;
               #TrFlowRefComp := #IOuMouldEditor_HMI.sSelected.sPS.arFlow[#RefComp];

               // Calculate ration out of flow rate
               FOR #TiLoop := 1 TO #TiComponentAmount DO
                   IF #TiLoop = #RefComp THEN
                       #IOuMouldEditor_HMI.sSelected.sPS.arRatio[#TiLoop] := 100.0;
                   ELSE
                       IF #TrFlowRefComp > 0 THEN
                           #IOuMouldEditor_HMI.sSelected.sPS.arRatio[#TiLoop] := #IOuMouldEditor_HMI.sSelected.sPS.arFlow[#TiLoop] * 100.0 / #TrFlowRefComp;
                       END_IF;
                   END_IF;
               END_FOR;
               //------------------------------------------------------------------------------------------------------------------------------------------------

               //  Value changed + Save data for the last cycle to recognize changes of the values
               //#IOuMouldEditor_HMI.sStatusBits.xValueChanged := TRUE;
               #SuMouldEditor_HMI := #IOuMouldEditor_HMI;
               // ----
               RETURN;
           END_IF;
       END_REGION
       //_________________________________________________________________________________    
       REGION Shot Time - changed
           FOR #TiLoop_PS := 1 TO #TiPartShotAmount DO
               IF #IOuMouldEditor_HMI.arShotSet[#TiLoop_PS].FoamingTime <> #SuMouldEditor_HMI.arShotSet[#TiLoop_PS].FoamingTime THEN
                   //  Calculation = 1 -> flow fixed
                   IF #IOuMouldEditor_HMI.sSelected.iCalculation = 1 THEN
                       #IOuMouldEditor_HMI.arShotSet[#TiLoop_PS].PartWeight := #IOuMouldEditor_HMI.arShotSet[#TiLoop_PS].FoamingTime * #IOuMouldEditor_HMI.sCalculatedValues.arTotalFlow[#TiLoop_PS];
                   END_IF;
                   // ----

                   //  Calculation = 2 -> weight fixed
                   IF #IOuMouldEditor_HMI.sSelected.iCalculation = 2 THEN
                       IF #IOuMouldEditor_HMI.arShotSet[#TiLoop_PS].FoamingTime > 0 THEN
                           #IOuMouldEditor_HMI.sCalculatedValues.arTotalFlow[#TiLoop_PS] := #IOuMouldEditor_HMI.arShotSet[#TiLoop_PS].PartWeight / #IOuMouldEditor_HMI.arShotSet[#TiLoop_PS].FoamingTime;

                           // SumRatio
                           #OUTrSumRatio := 0;

                           FOR #TiLoop_Ratio := 1 TO #TiComponentAmount DO
                               #OUTrSumRatio := #OUTrSumRatio + #IOuMouldEditor_HMI.sSelected.sPS.arRatio[#TiLoop_Ratio];
                           END_FOR;

                           FOR #TiLoop := 1 TO #TiComponentAmount DO
                               // only change single flow rates!                      
                               #IOuMouldEditor_HMI.sSelected.sPS.arFlow[#TiLoop] := #IOuMouldEditor_HMI.sCalculatedValues.arTotalFlow[#IOuMouldEditor_HMI.sSelected.sPS.iPS] /
                               #OUTrSumRatio * #IOuMouldEditor_HMI.sSelected.sPS.arRatio[#TiLoop];
                               #IOuMouldEditor_HMI.arShotSet[#IOuMouldEditor_HMI.sSelected.sPS.iPS].Flow[#TiLoop] := #IOuMouldEditor_HMI.sSelected.sPS.arFlow[#TiLoop];
                           END_FOR;
                       ELSE
                           #IOuMouldEditor_HMI.sCalculatedValues.arTotalFlow[#TiLoop_PS] := 0;
                           FOR #TiLoop := 1 TO #TiComponentAmount DO
                               #IOuMouldEditor_HMI.sSelected.sPS.arFlow[#TiLoop] := 0;
                               #IOuMouldEditor_HMI.arShotSet[#IOuMouldEditor_HMI.sSelected.sPS.iPS].Flow[#TiLoop] := #IOuMouldEditor_HMI.sSelected.sPS.arFlow[#TiLoop];
                           END_FOR;
                       END_IF;

                   END_IF;
                   // ----

                   //  Value changed + Save data for the last cycle to recognize changes of the values
                   #IOuMouldEditor_HMI.sStatusBits.xValueChanged := TRUE;
                   #SuMouldEditor_HMI := #IOuMouldEditor_HMI;
                   EXIT;
                   // ----

               END_IF
               ;
           END_FOR;
       END_REGION
       //_________________________________________________________________________________    
       REGION Total flow - changed
           FOR #TiLoop_PS := 1 TO #TiPartShotAmount DO
               IF #IOuMouldEditor_HMI.sCalculatedValues.arTotalFlow[#TiLoop_PS] <> #SuMouldEditor_HMI.sCalculatedValues.arTotalFlow[#TiLoop_PS] THEN
                   // SumRatio
                   #OUTrSumRatio := 0;

                   FOR #TiLoop_Ratio := 1 TO #TiComponentAmount DO
                       #OUTrSumRatio := #OUTrSumRatio + #IOuMouldEditor_HMI.sSelected.sPS.arRatio[#TiLoop_Ratio];
                   END_FOR;

                   FOR #TiLoop := 1 TO #TiComponentAmount DO
                       IF #IOuMouldEditor_HMI.sCalculatedValues.arTotalFlow[#TiLoop_PS] > 0 THEN
                           // only change single flow rates!                      
                           #IOuMouldEditor_HMI.sSelected.sPS.arFlow[#TiLoop] := #IOuMouldEditor_HMI.sCalculatedValues.arTotalFlow[#IOuMouldEditor_HMI.sSelected.sPS.iPS] /
                           #OUTrSumRatio * #IOuMouldEditor_HMI.sSelected.sPS.arRatio[#TiLoop];
                       ELSE
                           #IOuMouldEditor_HMI.sSelected.sPS.arFlow[#TiLoop] := 0;
                       END_IF;
                       #IOuMouldEditor_HMI.arShotSet[#IOuMouldEditor_HMI.sSelected.sPS.iPS].Flow[#TiLoop] := #IOuMouldEditor_HMI.sSelected.sPS.arFlow[#TiLoop];
                   END_FOR;

                   //  Calculation = 0 -> shot time fixed
                   IF #IOuMouldEditor_HMI.sSelected.iCalculation = 0 THEN
                       #IOuMouldEditor_HMI.arShotSet[#TiLoop_PS].PartWeight := #IOuMouldEditor_HMI.sCalculatedValues.arTotalFlow[#TiLoop_PS] * #IOuMouldEditor_HMI.arShotSet[#TiLoop_PS].FoamingTime;
                   END_IF;
                   // ----

                   //  Calculation = 2 -> weight fixed
                   IF #IOuMouldEditor_HMI.sSelected.iCalculation = 2 THEN
                       IF #IOuMouldEditor_HMI.sCalculatedValues.arTotalFlow[#TiLoop_PS] > 0 THEN
                           #IOuMouldEditor_HMI.arShotSet[#TiLoop_PS].FoamingTime := #IOuMouldEditor_HMI.arShotSet[#TiLoop_PS].PartWeight / #IOuMouldEditor_HMI.sCalculatedValues.arTotalFlow[#TiLoop_PS];
                       ELSE
                           #IOuMouldEditor_HMI.arShotSet[#TiLoop_PS].FoamingTime := 0;
                       END_IF;
                   END_IF;
                   // ----

                   //  Value changed + Save data for the last cycle to recognize changes of the values
                   #IOuMouldEditor_HMI.sStatusBits.xValueChanged := TRUE;
                   #SuMouldEditor_HMI := #IOuMouldEditor_HMI;
                   EXIT;
                   // ----

               END_IF
               ;
           END_FOR;
       END_REGION
       //_________________________________________________________________________________    
       REGION Total weight - changed
           FOR #TiLoop_PS := 1 TO #TiPartShotAmount DO
               IF #IOuMouldEditor_HMI.arShotSet[#TiLoop_PS].PartWeight <> #SuMouldEditor_HMI.arShotSet[#TiLoop_PS].PartWeight THEN

                   //  Calculation = 0 -> shot time fixed
                   IF #IOuMouldEditor_HMI.sSelected.iCalculation = 0 THEN
                       IF #IOuMouldEditor_HMI.arShotSet[#TiLoop_PS].PartWeight > 0 THEN
                           #IOuMouldEditor_HMI.sCalculatedValues.arTotalFlow[#TiLoop_PS] := #IOuMouldEditor_HMI.arShotSet[#TiLoop_PS].PartWeight / #IOuMouldEditor_HMI.arShotSet[#TiLoop_PS].FoamingTime;

                           // SumRatio
                           #OUTrSumRatio := 0;

                           FOR #TiLoop_Ratio := 1 TO #TiComponentAmount DO
                               #OUTrSumRatio := #OUTrSumRatio + #IOuMouldEditor_HMI.sSelected.sPS.arRatio[#TiLoop_Ratio];
                           END_FOR;

                           FOR #TiLoop_Flow := 1 TO #TiComponentAmount DO

                               #IOuMouldEditor_HMI.sSelected.sPS.arFlow[#TiLoop_Flow] := #IOuMouldEditor_HMI.sCalculatedValues.arTotalFlow[#IOuMouldEditor_HMI.sSelected.sPS.iPS] /
                               #OUTrSumRatio * #IOuMouldEditor_HMI.sSelected.sPS.arRatio[#TiLoop_Flow];
                               #IOuMouldEditor_HMI.arShotSet[#IOuMouldEditor_HMI.sSelected.sPS.iPS].Flow[#TiLoop_Flow] := #IOuMouldEditor_HMI.sSelected.sPS.arFlow[#TiLoop_Flow];
                           END_FOR;
                       ELSE
                           #IOuMouldEditor_HMI.sCalculatedValues.arTotalFlow[#TiLoop_PS] := 0;
                           FOR #TiLoop_Flow := 1 TO #TiComponentAmount DO
                               #IOuMouldEditor_HMI.sSelected.sPS.arFlow[#TiLoop_Flow] := 0;
                               #IOuMouldEditor_HMI.arShotSet[#IOuMouldEditor_HMI.sSelected.sPS.iPS].Flow[#TiLoop_Flow] := #IOuMouldEditor_HMI.sSelected.sPS.arFlow[#TiLoop_Flow];
                           END_FOR;
                       END_IF;

                   END_IF;
                   // ----

                   //  Calculation = 1 -> flow fixed
                   IF #IOuMouldEditor_HMI.sSelected.iCalculation = 1 THEN
                       IF #IOuMouldEditor_HMI.arShotSet[#TiLoop_PS].PartWeight > 0 THEN
                           #IOuMouldEditor_HMI.arShotSet[#TiLoop_PS].FoamingTime := #IOuMouldEditor_HMI.arShotSet[#TiLoop_PS].PartWeight / #IOuMouldEditor_HMI.sCalculatedValues.arTotalFlow[#TiLoop_PS];
                       ELSE
                           #IOuMouldEditor_HMI.arShotSet[#TiLoop_PS].FoamingTime := 0;
                       END_IF;
                   END_IF;
                   // ----

                   //  Value changed + Save data for the last cycle to recognize changes of the values
                   #IOuMouldEditor_HMI.sStatusBits.xValueChanged := TRUE;
                   #SuMouldEditor_HMI := #IOuMouldEditor_HMI;
                   EXIT;
                   // ----

               END_IF;
           END_FOR;
       END_REGION
       //_________________________________________________________________________________    
       REGION Flow - changed
           FOR #TiLoop := 1 TO #TiComponentAmount DO
               IF #IOuMouldEditor_HMI.sSelected.sPS.arFlow[#TiLoop] <> #SuMouldEditor_HMI.sSelected.sPS.arFlow[#TiLoop] THEN
                   // If Refcomp flowrate change --> change all mixing ratios on all other components
                   // if any other flowrate change --> change only this mixing ratio
                   // change total flow always